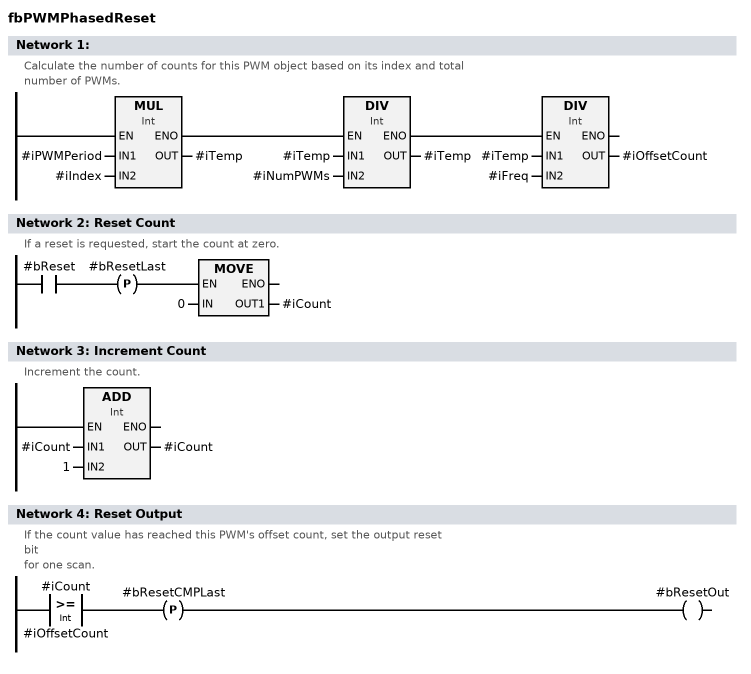
   RUNG wire#powerrail
      { S7_Templates := "SrcType := Int"; S7_GenerateENO := "TRUE" } Mul(in1 := #iPWMPeriod, in2 := #iIndex, out => #iTemp)
      { S7_Templates := "SrcType := Int"; S7_GenerateENO := "TRUE" } Div(in1 := #iTemp, in2 := #iNumPWMs, out => #iTemp)
      { S7_Templates := "SrcType := Int"; S7_GenerateENO := "TRUE" } Div(in1 := #iTemp, in2 := #iFreq, out => #iOffsetCount)
   END_RUNG
   // the same network as SCL:
   // ENO of a box is taken as its EN; it also drops when the box reports an error
   #iTemp := #iPWMPeriod * #iIndex;
   #iTemp := #iTemp / #iNumPWMs;
   #iOffsetCount := #iTemp / #iFreq;
END_REGION

REGION Network 2: Reset Count
   // If a reset is requested, start the count at zero.
   RUNG wire#powerrail
      Contact( #bReset )
      P_Trig( #bResetLast )
      { S7_GenerateENO := "TRUE" } Move(in := 0, out1 => #iCount)
   END_RUNG
   // the same network as SCL:
   #_w1 := #bReset AND NOT #bResetLast;   // rising edge
   #bResetLast := #bReset;
   IF #_w1 THEN #iCount := 0; END_IF;
END_REGION

REGION Network 3: Increment Count
   // Increment the count.
   RUNG wire#powerrail
      { S7_Templates := "SrcType := Int"; S7_GenerateENO := "TRUE" } Add(in1 := #iCount, in2 := 1, out => #iCount)
   END_RUNG
   // the same network as SCL:
   #iCount := #iCount + 1;
END_REGION

REGION Network 4: Reset Output
   // If the count value has reached this PWM's offset count, set the output reset 
   // bit 
   // for one scan.
   RUNG wire#powerrail
      { S7_Templates := "SrcType := Int" } GE_Contact(in1 := #iCount, in2 := #iOffsetCount)
      P_Trig( #bResetCMPLast )
      Coil( #bResetOut )
   END_RUNG
   // the same network as SCL:
   #_w1 := #iCount >= #iOffsetCount;
   #_w2 := #_w1 AND NOT #bResetCMPLast;   // rising edge
   #bResetCMPLast := #_w1;
   #bResetOut := #_w2;
END_REGION
END_FUNCTION_BLOCK

FUNCTION_BLOCK "fbRateCalc"   // FB170, LAD
TITLE = Calculate flow rate based on weight change
{ S7_Optimized_Access := 'FALSE' }
AUTHOR : DMC
FAMILY : RateCtrl
VERSION : 1.0
BEGIN

REGION Network 1: Sampling timer
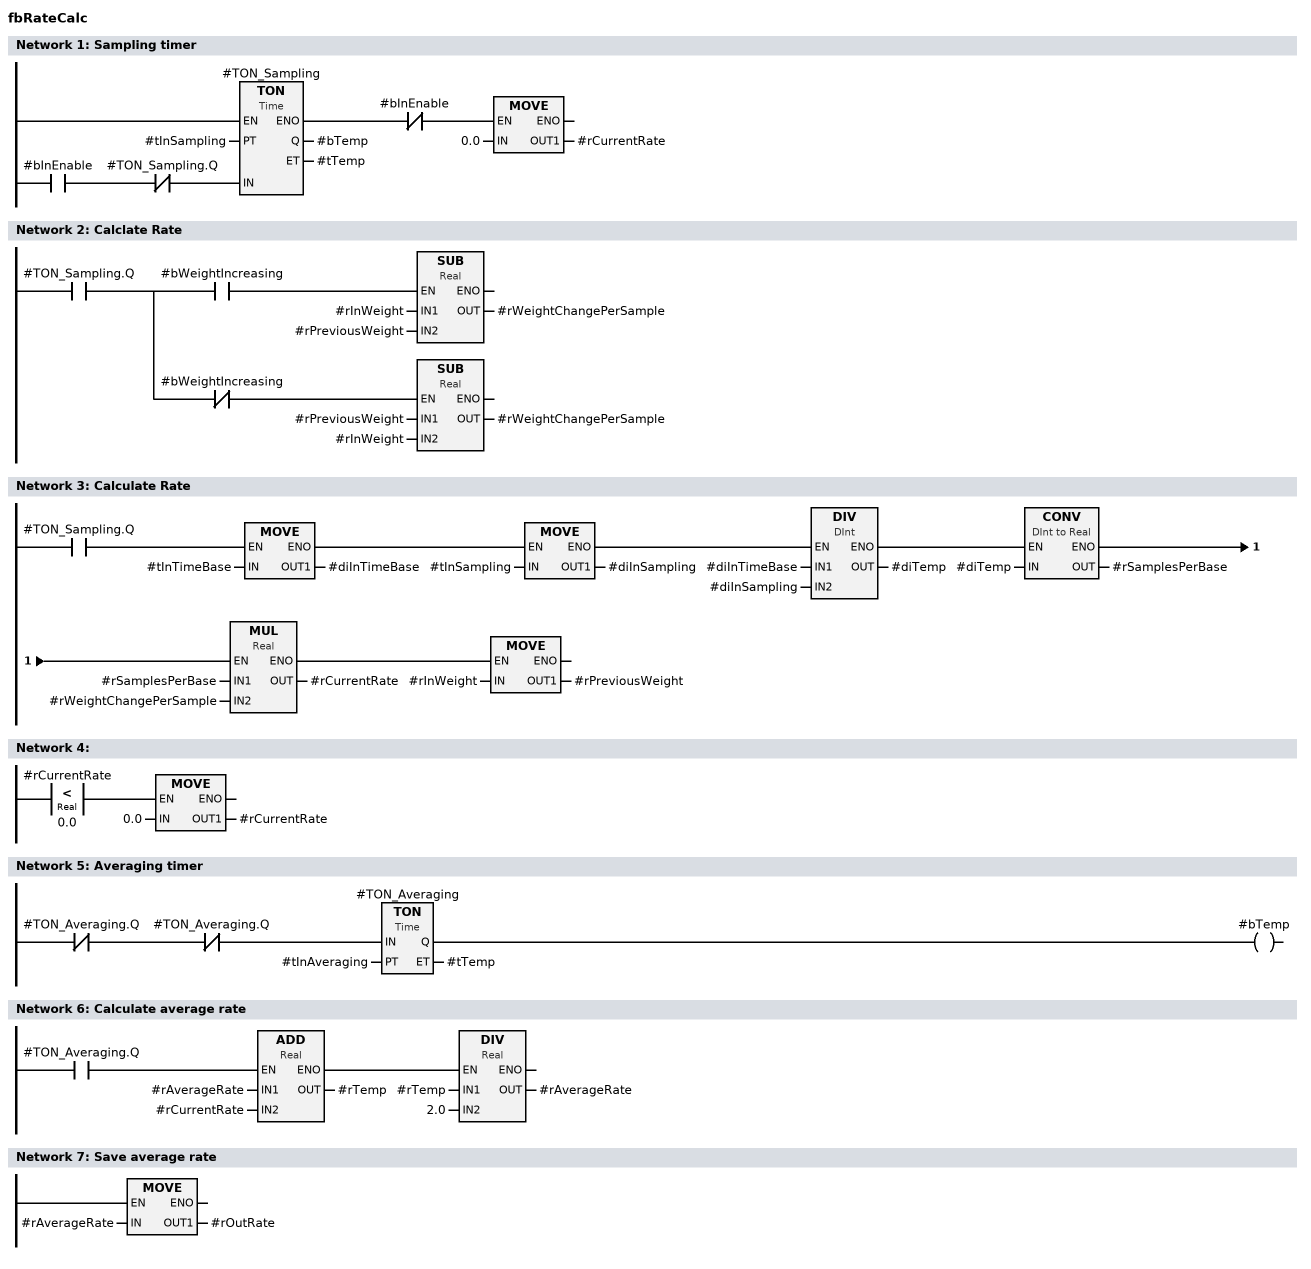
   // ENO of a box is taken as its EN; it also drops when the box reports an error
   #TON_Sampling.TON(pt := #tInSampling, in := #bInEnable AND NOT #TON_Sampling.Q, q => #bTemp, et => #tTemp);
   IF NOT #bInEnable THEN #rCurrentRate := 0.0; END_IF;
END_REGION

REGION Network 2: Calclate Rate
   RUNG wire#powerrail
      Contact( #TON_Sampling.Q )
      wire#w1
      Contact( #bWeightIncreasing )
      { S7_Templates := "SrcType := Real"; S7_GenerateENO := "TRUE" } Sub(in1 := #rInWeight, in2 := #rPreviousWeight, out => #rWeightChangePerSample)
   END_RUNG
   RUNG wire#w1
      I_Contact( #bWeightIncreasing )
      { S7_Templates := "SrcType := Real"; S7_GenerateENO := "TRUE" } Sub(in1 := #rPreviousWeight, in2 := #rInWeight, out => #rWeightChangePerSample)
   END_RUNG
   // the same network as SCL:
   IF #TON_Sampling.Q AND #bWeightIncreasing THEN
       #rWeightChangePerSample := #rInWeight - #rPreviousWeight;
   END_IF;
   IF #TON_Sampling.Q AND NOT #bWeightIncreasing THEN
       #rWeightChangePerSample := #rPreviousWeight - #rInWeight;
   END_IF;
END_REGION

REGION Network 3: Calculate Rate
   RUNG wire#powerrail
      Contact( #TON_Sampling.Q )
      { S7_GenerateENO := "TRUE" } Move(in := #tInTimeBase, out1 => #diInTimeBase)
      { S7_GenerateENO := "TRUE" } Move(in := #tInSampling, out1 => #diInSampling)
      { S7_Templates := "SrcType := DInt"; S7_GenerateENO := "TRUE" } Div(in1 := #diInTimeBase, in2 := #diInSampling, out => #diTemp)
      { S7_Templates := "[SrcType := DInt, DestType := Real]"; S7_GenerateENO := "TRUE" } Convert(in := #diTemp, out => #rSamplesPerBase)
      { S7_Templates := "SrcType := Real"; S7_GenerateENO := "TRUE" } Mul(in1 := #rSamplesPerBase, in2 := #rWeightChangePerSample, out => #rCurrentRate)
      { S7_GenerateENO := "TRUE" } Move(in := #rInWeight, out1 => #rPreviousWeight)
   END_RUNG
   // the same network as SCL:
   // ENO of a box is taken as its EN; it also drops when the box reports an error
   IF #TON_Sampling.Q THEN
       #diInTimeBase := #tInTimeBase;
       #diInSampling := #tInSampling;
       #diTemp := #diInTimeBase / #diInSampling;
       #rSamplesPerBase := DINT_TO_REAL(#diTemp);
       #rCurrentRate := #rSamplesPerBase * #rWeightChangePerSample;
       #rPreviousWeight := #rInWeight;
   END_IF;
END_REGION

REGION Network 4
   RUNG wire#powerrail
      { S7_Templates := "SrcType := Real" } LT_Contact(in1 := #rCurrentRate, in2 := 0.0)
      { S7_GenerateENO := "TRUE" } Move(in := 0.0, out1 => #rCurrentRate)
   END_RUNG
   // the same network as SCL:
   IF #rCurrentRate < 0.0 THEN #rCurrentRate := 0.0; END_IF;
END_REGION

REGION Network 5: Averaging timer
   #TON_Averaging.TON(pt := #tInAveraging, in := NOT #TON_Averaging.Q AND NOT #TON_Averaging.Q, et => #tTemp);
   #bTemp := #TON_Averaging.q;
END_REGION

REGION Network 6: Calculate average rate
   RUNG wire#powerrail
      Contact( #TON_Averaging.Q )
      { S7_Templates := "SrcType := Real"; S7_GenerateENO := "TRUE" } Add(in1 := #rAverageRate, in2 := #rCurrentRate, out => #rTemp)
      { S7_Templates := "SrcType := Real"; S7_GenerateENO := "TRUE" } Div(in1 := #rTemp, in2 := 2.0, out => #rAverageRate)
   END_RUNG
   // the same network as SCL:
   // ENO of a box is taken as its EN; it also drops when the box reports an error
   IF #TON_Averaging.Q THEN
       #rTemp := #rAverageRate + #rCurrentRate;
       #rAverageRate := #rTemp / 2.0;
   END_IF;
END_REGION

REGION Network 7: Save average rate
   RUNG wire#powerrail
      { S7_GenerateENO := "TRUE" } Move(in := #rAverageRate, out1 => #rOutRate)
   END_RUNG
   // the same network as SCL:
   #rOutRate := #rAverageRate;
END_REGION

REGION Network 8 (STL): Set ENO bit

         SET;
         SAVE;
END_REGION
END_FUNCTION_BLOCK

FUNCTION_BLOCK "fbPulser"   // FB173, LAD
{ S7_Optimized_Access := 'FALSE' }
VERSION : 0.1
BEGIN

REGION Network 1 (STL)
   // added on time and off time to obtain a period
         L     #tIN_TIME_ON;
         L     #tIN_TIME_OFF;
         +D;
         T     #tTIME_TOTAL;
END_REGION

REGION Network 2 (STL)
   // Verify that tInTIME_ON and OFF are bigger than 0

         L     #tIN_TIME_ON;
         L     T#0MS;
         ==D;
         =     #bOn_0;

         L     #tIN_TIME_OFF;
         L     T#0MS;
         ==D;
         =     #bOff_0;
END_REGION

REGION Network 3
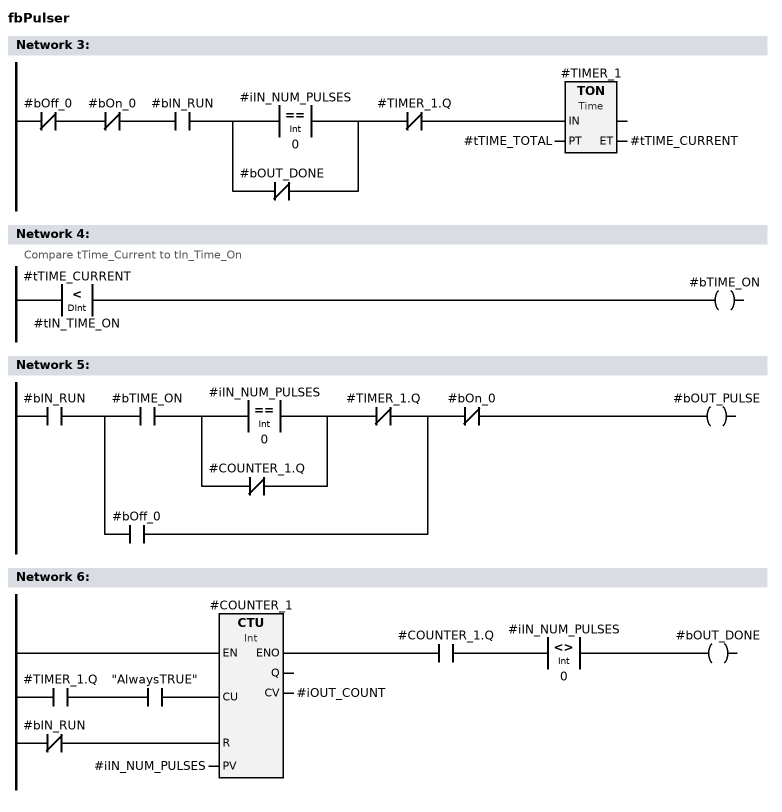
   #TIMER_1.TON(pt := #tTIME_TOTAL,
                in := NOT #bOff_0 AND NOT #bOn_0 AND #bIN_RUN AND ((#iIN_NUM_PULSES = 0) OR NOT #bOUT_DONE) AND NOT #TIMER_1.Q,
                et => #tTIME_CURRENT);
END_REGION

REGION Network 4
   // Compare tTime_Current to tIn_Time_On
   RUNG wire#powerrail
      { S7_Templates := "SrcType := DInt" } LT_Contact(in1 := #tTIME_CURRENT, in2 := #tIN_TIME_ON)
      Coil( #bTIME_ON )
   END_RUNG
   // the same network as SCL:
   #bTIME_ON := #tTIME_CURRENT < #tIN_TIME_ON;
END_REGION

REGION Network 5
   #bOUT_PULSE := #bIN_RUN AND ((#bTIME_ON AND ((#iIN_NUM_PULSES = 0) OR NOT #COUNTER_1.Q) AND NOT #TIMER_1.Q) OR #bOff_0) AND NOT #bOn_0;
END_REGION

REGION Network 6
   // ENO of a box is taken as its EN; it also drops when the box reports an error
   #COUNTER_1.CTU(CU := #TIMER_1.Q AND "AlwaysTRUE",
                  R := NOT #bIN_RUN,
                  PV := #iIN_NUM_PULSES,
                  CV => #iOUT_COUNT);
   #bOUT_DONE := #COUNTER_1.Q AND (#iIN_NUM_PULSES <> 0);
END_REGION
END_FUNCTION_BLOCK

FUNCTION_BLOCK "fbRunningAverage"   // FB196, SCL
TITLE = Running average calculation
{ S7_Optimized_Access := 'FALSE' }
AUTHOR : DMC
VERSION : 1.10
// 2012-05-23 DMC-BC: Added min/max
BEGIN


   // Shift history array left by 1
   #iTemp:=BLKMOV(SRCBLK := #ValueHistoryFrom.Sub, DSTBLK => #Sub);
   #iTemp:=BLKMOV(SRCBLK := #Sub, DSTBLK => #ValueHistoryTo.Sub);

   // Add new value
   #ValueHistory[1] := #rInValue;

   IF #iInBufferSize > 1 THEN

       // Limit buffer size to the size of the array
       IF #iInBufferSize <= #ciSize THEN
           #iOutBufferSize := #iInBufferSize;
           #bOutError := false;
       ELSE
           #iOutBufferSize := #ciSize; 
           #bOutError := true;
       END_IF;

       // Cycle throough the array
       #rSum := 0.0;
       #rMax := -3.402822E+38;
       #rMin := 3.402822E+38;
       FOR #i:=1 TO #iOutBufferSize BY 1 DO  

           // Min/max logic
           IF #ValueHistory[#i] > #rMax THEN
               #rMax := #ValueHistory[#i];
           END_IF;                
           IF #ValueHistory[#i] < #rMin THEN
               #rMin := #ValueHistory[#i];
           END_IF;

           // Calcualte sum
           #rSum := #rSum + #ValueHistory[#i];
       END_FOR;

       // Calculate average
       #rOutAverage := #rSum /(DINT_TO_REAL(#iOutBufferSize));
       #rOutMin := #rMin;
       #rOutMax := #rMax;
   ELSE
       // Buffer size is 1 - no averaging
       #iOutBufferSize := 1;
       #rOutAverage := #rInValue;
       #rOutMin := #rInValue;
       #rOutMax := #rInValue;
   END_IF;

   ENO:=true;
END_FUNCTION_BLOCK

FUNCTION_BLOCK "fbRetentiveTimer"   // FB1011, LAD
TITLE = Retentive Timer Block
{ S7_Optimized_Access := 'FALSE' }
AUTHOR : DMC
FAMILY : LowLevel
VERSION : 0.1
// //  This is a retentive count-up timer.
// //  IN makes it count.  It does not reset when IN is off.
// //  RESET resets the time to 0.  
// //  bInPT is the time setpoint.
// //  bOutEnabled is true when the time has the setpoint
// //  bOutET is the elapsed time.
   VAR_TEMP   // added for the SCL form of the ladder/FBD networks
      _w1 : Bool;
   END_VAR
BEGIN

REGION Network 1: Keep resetting internal time while not counting
   // IF (NOT IN) THEN
   //     tInternalTime := tInternalTime + Timer1.ET;
   // END_IF;
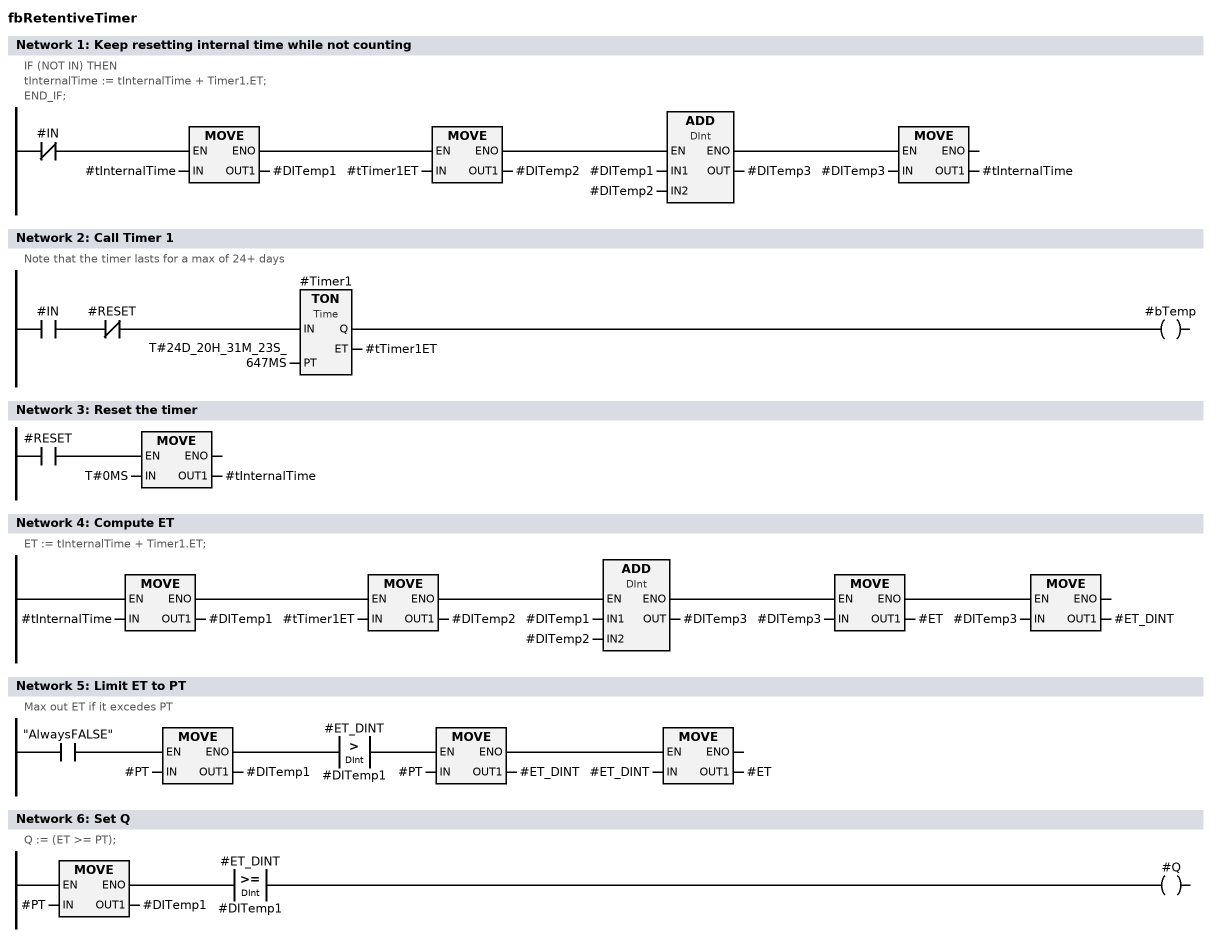
   RUNG wire#powerrail
      I_Contact( #IN )
      { S7_GenerateENO := "TRUE" } Move(in := #tInternalTime, out1 => #DITemp1)
      { S7_GenerateENO := "TRUE" } Move(in := #tTimer1ET, out1 => #DITemp2)
      { S7_Templates := "SrcType := DInt"; S7_GenerateENO := "TRUE" } Add(in1 := #DITemp1, in2 := #DITemp2, out => #DITemp3)
      { S7_GenerateENO := "TRUE" } Move(in := #DITemp3, out1 => #tInternalTime)
   END_RUNG
   // the same network as SCL:
   // ENO of a box is taken as its EN; it also drops when the box reports an error
   IF NOT #IN THEN
       #DITemp1 := #tInternalTime;
       #DITemp2 := #tTimer1ET;
       #DITemp3 := #DITemp1 + #DITemp2;
       #tInternalTime := #DITemp3;
   END_IF;
END_REGION

REGION Network 2: Call Timer 1
   // Note that the timer lasts for a max of 24+ days
   #Timer1.TON(IN := #IN AND NOT #RESET, PT := T#24D_20H_31M_23S_647MS, ET => #tTimer1ET);
   #bTemp := #Timer1.Q;
END_REGION

REGION Network 3: Reset the timer
   RUNG wire#powerrail
      Contact( #RESET )
      { S7_GenerateENO := "TRUE" } Move(in := T#0MS, out1 => #tInternalTime)
   END_RUNG
   // the same network as SCL:
   IF #RESET THEN #tInternalTime := T#0MS; END_IF;
END_REGION

REGION Network 4: Compute ET
   // ET := tInternalTime + Timer1.ET;
   RUNG wire#powerrail
      { S7_GenerateENO := "TRUE" } Move(in := #tInternalTime, out1 => #DITemp1)
      { S7_GenerateENO := "TRUE" } Move(in := #tTimer1ET, out1 => #DITemp2)
      { S7_Templates := "SrcType := DInt"; S7_GenerateENO := "TRUE" } Add(in1 := #DITemp1, in2 := #DITemp2, out => #DITemp3)
      { S7_GenerateENO := "TRUE" } Move(in := #DITemp3, out1 => #ET)
      { S7_GenerateENO := "TRUE" } Move(in := #DITemp3, out1 => #ET_DINT)
   END_RUNG
   // the same network as SCL:
   // ENO of a box is taken as its EN; it also drops when the box reports an error
   #DITemp1 := #tInternalTime;
   #DITemp2 := #tTimer1ET;
   #DITemp3 := #DITemp1 + #DITemp2;
   #ET := #DITemp3;
   #ET_DINT := #DITemp3;
END_REGION

REGION Network 5: Limit ET to PT
   // Max out ET if it excedes PT
   RUNG wire#powerrail
      Contact( "AlwaysFALSE" )
      { S7_GenerateENO := "TRUE" } Move(in := #PT, out1 => #DITemp1)
      { S7_Templates := "SrcType := DInt" } GT_Contact(in1 := #ET_DINT, in2 := #DITemp1)
      { S7_GenerateENO := "TRUE" } Move(in := #PT, out1 => #ET_DINT)
      { S7_GenerateENO := "TRUE" } Move(in := #ET_DINT, out1 => #ET)
   END_RUNG
   // the same network as SCL:
   // ENO of a box is taken as its EN; it also drops when the box reports an error
   IF "AlwaysFALSE" THEN #DITemp1 := #PT; END_IF;
   #_w1 := "AlwaysFALSE" AND (#ET_DINT > #DITemp1);
   IF #_w1 THEN
       #ET_DINT := #PT;
       #ET := #ET_DINT;
   END_IF;
END_REGION

REGION Network 6: Set Q
   // Q := (ET >= PT);
   RUNG wire#powerrail
      { S7_GenerateENO := "TRUE" } Move(in := #PT, out1 => #DITemp1)
      { S7_Templates := "SrcType := DInt" } GE_Contact(in1 := #ET_DINT, in2 := #DITemp1)
      Coil( #Q )
   END_RUNG
   // the same network as SCL:
   // ENO of a box is taken as its EN; it also drops when the box reports an error
   #DITemp1 := #PT;
   #Q := #ET_DINT >= #DITemp1;
END_REGION
END_FUNCTION_BLOCK

FUNCTION_BLOCK "fbRetentiveTimer"   // FB1940, LAD
TITLE = Retentive Timer Block
{ S7_Optimized_Access := 'FALSE' }
AUTHOR : DMC
FAMILY : LowLevel
VERSION : 0.1
// //  This is a retentive count-up timer.
// //  IN makes it count.  It does not reset when IN is off.
// //  RESET resets the time to 0.  
// //  PT is the time setpoint.
// //  Q is true when the time has the setpoint
// //  ET is the elapsed time (ms)
   VAR_TEMP   // added for the SCL form of the ladder/FBD networks
      _w1 : Bool;
      _w2 : Bool;
   END_VAR
BEGIN

REGION Network 1: Keep resetting internal time while not counting
   // IF (NOT IN) THEN
   //     tInternalTime := tInternalTime + Timer1.ET;
   // END_IF;
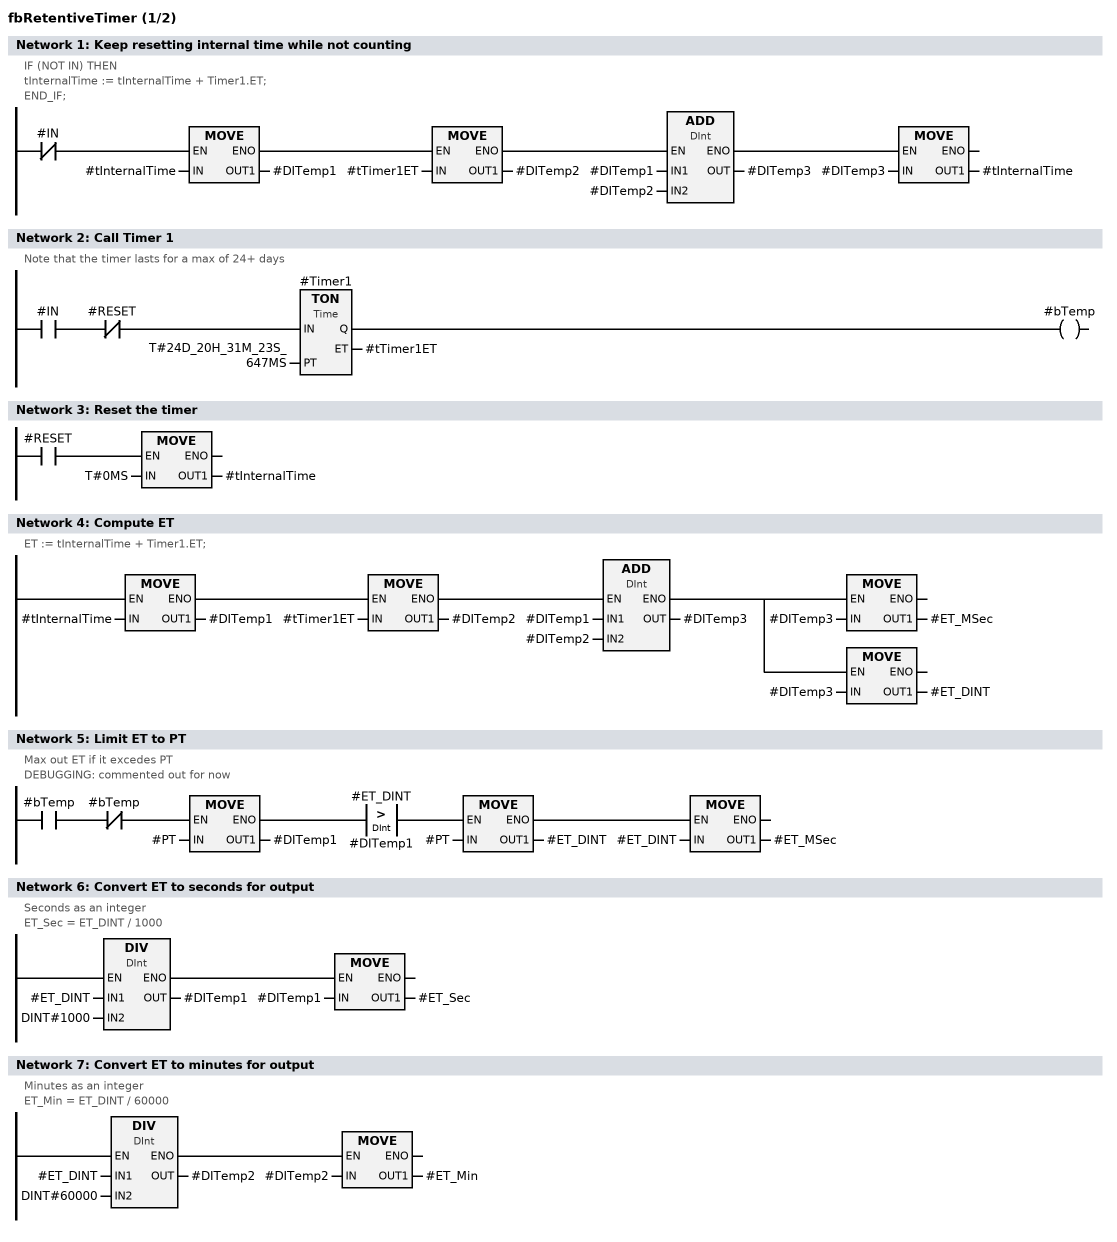
   RUNG wire#powerrail
      I_Contact( #IN )
      { S7_GenerateENO := "TRUE" } Move(in := #tInternalTime, out1 => #DITemp1)
      { S7_GenerateENO := "TRUE" } Move(in := #tTimer1ET, out1 => #DITemp2)
      { S7_Templates := "SrcType := DInt"; S7_GenerateENO := "TRUE" } Add(in1 := #DITemp1, in2 := #DITemp2, out => #DITemp3)
      { S7_GenerateENO := "TRUE" } Move(in := #DITemp3, out1 => #tInternalTime)
   END_RUNG
   // the same network as SCL:
   // ENO of a box is taken as its EN; it also drops when the box reports an error
   IF NOT #IN THEN
       #DITemp1 := #tInternalTime;
       #DITemp2 := #tTimer1ET;
       #DITemp3 := #DITemp1 + #DITemp2;
       #tInternalTime := #DITemp3;
   END_IF;
END_REGION

REGION Network 2: Call Timer 1
   // Note that the timer lasts for a max of 24+ days
   #Timer1.TON(pt := T#24D_20H_31M_23S_647MS, in := #IN AND NOT #RESET, et => #tTimer1ET);
   #bTemp := #Timer1.q;
END_REGION

REGION Network 3: Reset the timer
   RUNG wire#powerrail
      Contact( #RESET )
      { S7_GenerateENO := "TRUE" } Move(in := T#0MS, out1 => #tInternalTime)
   END_RUNG
   // the same network as SCL:
   IF #RESET THEN #tInternalTime := T#0MS; END_IF;
END_REGION

REGION Network 4: Compute ET
   // ET := tInternalTime + Timer1.ET;
   RUNG wire#powerrail
      { S7_GenerateENO := "TRUE" } Move(in := #tInternalTime, out1 => #DITemp1)
      { S7_GenerateENO := "TRUE" } Move(in := #tTimer1ET, out1 => #DITemp2)
      { S7_Templates := "SrcType := DInt"; S7_GenerateENO := "TRUE" } Add(in1 := #DITemp1, in2 := #DITemp2, out => #DITemp3)
      wire#w1
      { S7_GenerateENO := "TRUE" } Move(in := #DITemp3, out1 => #ET_MSec)
   END_RUNG
   RUNG wire#w1
      { S7_GenerateENO := "TRUE" } Move(in := #DITemp3, out1 => #ET_DINT)
   END_RUNG
   // the same network as SCL:
   // ENO of a box is taken as its EN; it also drops when the box reports an error
   #DITemp1 := #tInternalTime;
   #DITemp2 := #tTimer1ET;
   #DITemp3 := #DITemp1 + #DITemp2;
   #ET_MSec := #DITemp3;
   #ET_DINT := #DITemp3;
END_REGION

REGION Network 5: Limit ET to PT
   // Max out ET if it excedes PT
   // 
   // DEBUGGING: commented out for now
   RUNG wire#powerrail
      Contact( #bTemp )
      I_Contact( #bTemp )
      { S7_GenerateENO := "TRUE" } Move(in := #PT, out1 => #DITemp1)
      { S7_Templates := "SrcType := DInt" } GT_Contact(in1 := #ET_DINT, in2 := #DITemp1)
      { S7_GenerateENO := "TRUE" } Move(in := #PT, out1 => #ET_DINT)
      { S7_GenerateENO := "TRUE" } Move(in := #ET_DINT, out1 => #ET_MSec)
   END_RUNG
   // the same network as SCL:
   // ENO of a box is taken as its EN; it also drops when the box reports an error
   #_w1 := #bTemp AND NOT #bTemp;
   IF #_w1 THEN #DITemp1 := #PT; END_IF;
   #_w2 := #_w1 AND (#ET_DINT > #DITemp1);
   IF #_w2 THEN
       #ET_DINT := #PT;
       #ET_MSec := #ET_DINT;
   END_IF;
END_REGION

REGION Network 6: Convert ET to seconds for output
   // Seconds as an integer
   // ET_Sec = ET_DINT / 1000
   RUNG wire#powerrail
      { S7_Templates := "SrcType := DInt"; S7_GenerateENO := "TRUE" } Div(in1 := #ET_DINT, in2 := DINT#1000, out => #DITemp1)
      { S7_GenerateENO := "TRUE" } Move(in := #DITemp1, out1 => #ET_Sec)
   END_RUNG
   // the same network as SCL:
   // ENO of a box is taken as its EN; it also drops when the box reports an error
   #DITemp1 := #ET_DINT / DINT#1000;
   #ET_Sec := #DITemp1;
END_REGION

REGION Network 7: Convert ET to minutes for output
   // Minutes as an integer
   // ET_Min = ET_DINT / 60000
   RUNG wire#powerrail
      { S7_Templates := "SrcType := DInt"; S7_GenerateENO := "TRUE" } Div(in1 := #ET_DINT, in2 := DINT#60000, out => #DITemp2)
      { S7_GenerateENO := "TRUE" } Move(in := #DITemp2, out1 => #ET_Min)
   END_RUNG
   // the same network as SCL:
   // ENO of a box is taken as its EN; it also drops when the box reports an error
   #DITemp2 := #ET_DINT / DINT#60000;
   #ET_Min := #DITemp2;
END_REGION

REGION Network 8: Convert ET to hours for output
   // Hours as a real number (can show decimals of hours with 1/60 resolution)
   // ET_Hour = REAL(ET_Min) / 60.0
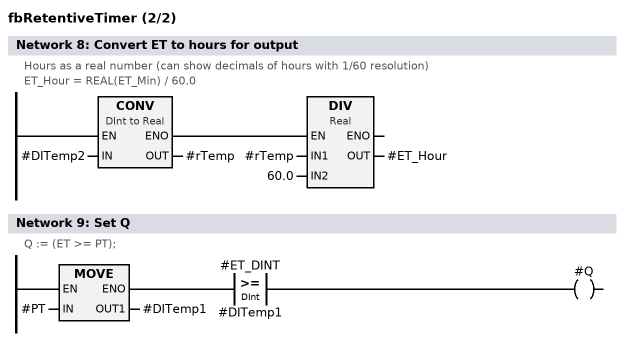
   RUNG wire#powerrail
      { S7_Templates := "[SrcType := DInt, DestType := Real]"; S7_GenerateENO := "TRUE" } Convert(in := #DITemp2, out => #rTemp)
      { S7_Templates := "SrcType := Real"; S7_GenerateENO := "TRUE" } Div(in1 := #rTemp, in2 := 60.0, out => #ET_Hour)
   END_RUNG
   // the same network as SCL:
   // ENO of a box is taken as its EN; it also drops when the box reports an error
   #rTemp := DINT_TO_REAL(#DITemp2);
   #ET_Hour := #rTemp / 60.0;
END_REGION

REGION Network 9: Set Q
   // Q := (ET >= PT);
   RUNG wire#powerrail
      { S7_GenerateENO := "TRUE" } Move(in := #PT, out1 => #DITemp1)
      { S7_Templates := "SrcType := DInt" } GE_Contact(in1 := #ET_DINT, in2 := #DITemp1)
      Coil( #Q )
   END_RUNG
   // the same network as SCL:
   // ENO of a box is taken as its EN; it also drops when the box reports an error
   #DITemp1 := #PT;
   #Q := #ET_DINT >= #DITemp1;
END_REGION

REGION Network 10 (STL): Set the Save Bit
         SET;
         SAVE;
END_REGION
END_FUNCTION_BLOCK

FUNCTION "fcTolerance" : Void   // FC1010, LAD
TITLE = Check if a value is in tolerance
{ S7_Optimized_Access := 'FALSE' }
AUTHOR : DMC
FAMILY : Recipe
VERSION : 0.1
BEGIN

REGION Network 1: Check value in tolerance
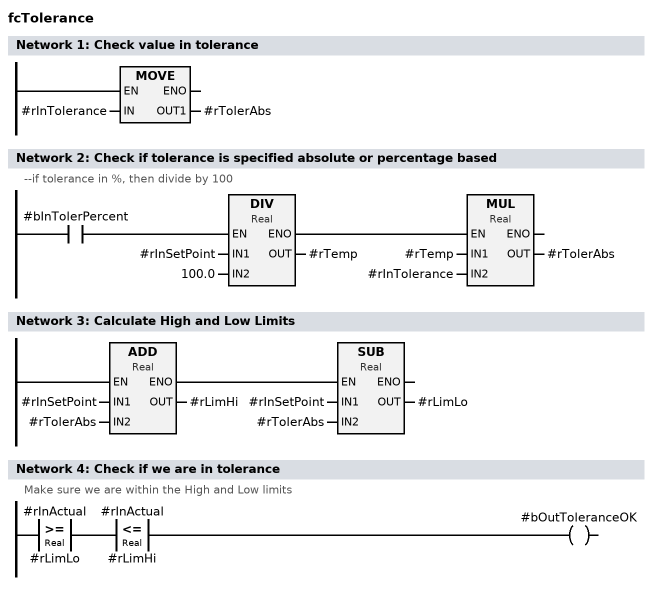
   RUNG wire#powerrail
      { S7_GenerateENO := "TRUE" } Move(in := #rInTolerance, out1 => #rTolerAbs)
   END_RUNG
   // the same network as SCL:
   #rTolerAbs := #rInTolerance;
END_REGION

REGION Network 2: Check if tolerance is specified absolute or percentage based
   // --if tolerance in %, then divide by 100
   RUNG wire#powerrail
      Contact( #bInTolerPercent )
      { S7_Templates := "SrcType := Real"; S7_GenerateENO := "TRUE" } Div(in1 := #rInSetPoint, in2 := 100.0, out => #rTemp)
      { S7_Templates := "SrcType := Real"; S7_GenerateENO := "TRUE" } Mul(in1 := #rTemp, in2 := #rInTolerance, out => #rTolerAbs)
   END_RUNG
   // the same network as SCL:
   // ENO of a box is taken as its EN; it also drops when the box reports an error
   IF #bInTolerPercent THEN
       #rTemp := #rInSetPoint / 100.0;
       #rTolerAbs := #rTemp * #rInTolerance;
   END_IF;
END_REGION

REGION Network 3: Calculate High and Low Limits
   RUNG wire#powerrail
      { S7_Templates := "SrcType := Real"; S7_GenerateENO := "TRUE" } Add(in1 := #rInSetPoint, in2 := #rTolerAbs, out => #rLimHi)
      { S7_Templates := "SrcType := Real"; S7_GenerateENO := "TRUE" } Sub(in1 := #rInSetPoint, in2 := #rTolerAbs, out => #rLimLo)
   END_RUNG
   // the same network as SCL:
   // ENO of a box is taken as its EN; it also drops when the box reports an error
   #rLimHi := #rInSetPoint + #rTolerAbs;
   #rLimLo := #rInSetPoint - #rTolerAbs;
END_REGION

REGION Network 4: Check if we are in tolerance
   // Make sure we are within the High and Low limits
   RUNG wire#powerrail
      { S7_Templates := "SrcType := Real" } GE_Contact(in1 := #rInActual, in2 := #rLimLo)
      { S7_Templates := "SrcType := Real" } LE_Contact(in1 := #rInActual, in2 := #rLimHi)
      Coil( #bOutToleranceOK )
   END_RUNG
   // the same network as SCL:
   #bOutToleranceOK := (#rInActual >= #rLimLo) AND (#rInActual <= #rLimHi);
END_REGION

REGION Network 5 (STL): Save RLO Bit
         SET;
         SAVE;
END_REGION
END_FUNCTION

FUNCTION "fcTolerance" : Void   // FC1010, LAD
TITLE = Check if a value is in tolerance
{ S7_Optimized_Access := 'FALSE' }
AUTHOR : DMC
FAMILY : Process
VERSION : 0.1
BEGIN

REGION Network 1: Check value in tolerance
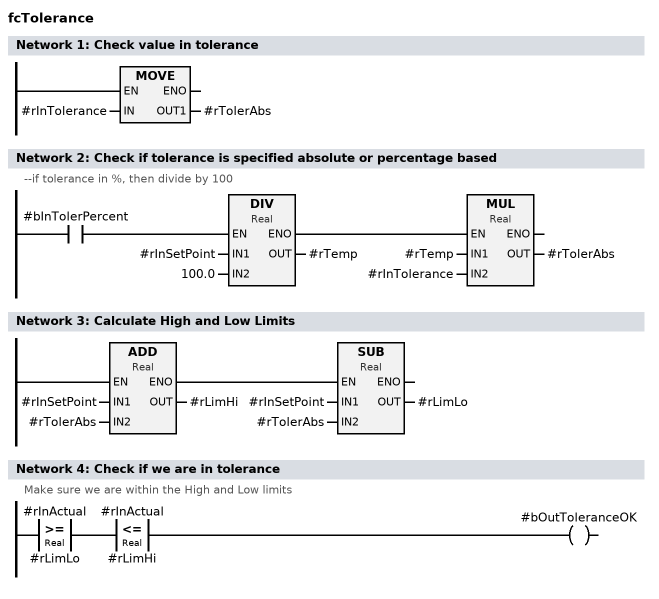
   RUNG wire#powerrail
      { S7_GenerateENO := "TRUE" } Move(in := #rInTolerance, out1 => #rTolerAbs)
   END_RUNG
   // the same network as SCL:
   #rTolerAbs := #rInTolerance;
END_REGION

REGION Network 2: Check if tolerance is specified absolute or percentage based
   // --if tolerance in %, then divide by 100
   RUNG wire#powerrail
      Contact( #bInTolerPercent )
      { S7_Templates := "SrcType := Real"; S7_GenerateENO := "TRUE" } Div(in1 := #rInSetPoint, in2 := 100.0, out => #rTemp)
      { S7_Templates := "SrcType := Real"; S7_GenerateENO := "TRUE" } Mul(in1 := #rTemp, in2 := #rInTolerance, out => #rTolerAbs)
   END_RUNG
   // the same network as SCL:
   // ENO of a box is taken as its EN; it also drops when the box reports an error
   IF #bInTolerPercent THEN
       #rTemp := #rInSetPoint / 100.0;
       #rTolerAbs := #rTemp * #rInTolerance;
   END_IF;
END_REGION

REGION Network 3: Calculate High and Low Limits
   RUNG wire#powerrail
      { S7_Templates := "SrcType := Real"; S7_GenerateENO := "TRUE" } Add(in1 := #rInSetPoint, in2 := #rTolerAbs, out => #rLimHi)
      { S7_Templates := "SrcType := Real"; S7_GenerateENO := "TRUE" } Sub(in1 := #rInSetPoint, in2 := #rTolerAbs, out => #rLimLo)
   END_RUNG
   // the same network as SCL:
   // ENO of a box is taken as its EN; it also drops when the box reports an error
   #rLimHi := #rInSetPoint + #rTolerAbs;
   #rLimLo := #rInSetPoint - #rTolerAbs;
END_REGION

REGION Network 4: Check if we are in tolerance
   // Make sure we are within the High and Low limits
   RUNG wire#powerrail
      { S7_Templates := "SrcType := Real" } GE_Contact(in1 := #rInActual, in2 := #rLimLo)
      { S7_Templates := "SrcType := Real" } LE_Contact(in1 := #rInActual, in2 := #rLimHi)
      Coil( #bOutToleranceOK )
   END_RUNG
   // the same network as SCL:
   #bOutToleranceOK := (#rInActual >= #rLimLo) AND (#rInActual <= #rLimHi);
END_REGION
END_FUNCTION

// ===== library: MasterCopy "Open Library" =====

VAR_GLOBAL   // PLC tag table "Open Library"
   "System_Byte" AT %MB1 : Byte;
   "FirstScan" AT %M1.0 : Bool;
   "DiagStatusUpdate" AT %M1.1 : Bool;
   "Clock_Byte" AT %MB0 : Byte;
   "Clock_10Hz" AT %M0.0 : Bool;
   "Clock_5Hz" AT %M0.1 : Bool;
   "Clock_2.5Hz" AT %M0.2 : Bool;
   "Clock_2Hz" AT %M0.3 : Bool;
   "Clock_1.25Hz" AT %M0.4 : Bool;
   "Clock_1Hz" AT %M0.5 : Bool;
   "Clock_0.625Hz" AT %M0.6 : Bool;
   "Clock_0.5Hz" AT %M0.7 : Bool;
   "AlwaysTRUE" AT %M1.2 : Bool;
   "AlwaysFALSE" AT %M1.3 : Bool;
END_VAR
